		IF SwitchIO.xLiftCylinderExtendInit THEN
		  	IF SwitchIO.xLiftCylinderRetractDetect THEN
		  		iStep:=4;
		  	END_IF;
		  	ELSE
		  	IF SwitchIO.xLiftCylinderExtendDetect THEN
				iStep:=4; 
		  	END_IF;
		END_IF;
		3:(*放行*)	
		ConveyorExitIO.iProductCategory:=ConveyorEntryIO.iProductCategory;
		ConveyorExitIO.iTaskID:=ConveyorEntryIO.iTaskID;
		ConveyorExitIO.diDesConveyor:=ConveyorEntryIO.diDesConveyor;
		SwitchIO.xExitBarCylinderRetract:=1;
		ConveyorExitIO.xPutInto:=0;
		iStep:=4;
		4:(*下料*)
		(*通过出料传输线下料*)
		IF SwitchIO.xExitEnable  AND m_xExitBarDelay AND NOT SwitchIO.xExitBarCylinderRetract  THEN		  
		  	ConveyorExitIO.xUnload:=1;
			ELSE
		  	ConveyorExitIO.xUnload:=0;
		END_IF;	
		(*通过进料传输线下料*)
		IF SwitchIO.xExitEnable  AND m_xExitBarDelay  AND SwitchIO.xExitBarCylinderRetract THEN		  
		  	ConveyorEntryIO.xUnload:=1;
			ELSE
		  	ConveyorEntryIO.xUnload:=0;
		END_IF;			    	
		IF (ConveyorExitIO.xEmpty OR ConveyorEntryIO.xEmpty) AND m_xExitBarDelay  THEN
		  	ConveyorExitIO.xPutInto:=1;
		  	ConveyorEntryIO.xPutInto:=1;
			iStep:=0; 
		END_IF;
	END_CASE;
	m_tonLiftCylinderDelay(IN:=NOT ConveyorEntryIO.xEmpty AND iStep=1 ,PT:= T#1S ,Q:= m_xLiftCylinderDelay ,ET:=m_tLiftCylinderDelay );
	m_tonExitBarDelay(IN:=iStep=4 ,PT:= T#1s ,Q:= m_xExitBarDelay ,ET:= m_tExitBarDelay);
END_IF;
(*复位程序*)
IF (g_xResetSingle AND  (g_diDeviceIDSelect=ConveyorEntryIO.diDeviceID OR g_diDeviceIDSelect=ConveyorExitIO.diDeviceID))
	OR LDP(TRUE,SwitchIO.xLiftCylinderExtendInit) 
	OR LDF(TRUE,SwitchIO.xLiftCylinderExtendInit) 
	OR LDP(TRUE,SwitchIO.xPutInto)  THEN
	ConveyorEntryIO.xPutInto:=1;
	ConveyorExitIO.xPutInto:=1;
	iStep:=0;
END_IF;

IF g_xManual  THEN
	iStep:=0;
	ConveyorEntryIO.xLoad:=0;
    ConveyorEntryIO.xUnload:=0;
	ConveyorEntryIO.xPutInto:=0;
	ConveyorExitIO.xLoad:=0;
	ConveyorExitIo.xUnload:=0;
	ConveyorExitIO.xPutInto:=0;
	SwitchIO.xEntryBarCylinderRetract:=0;
	SwitchIO.xExitBarCylinderRetract:=0;
	IF SwitchIO.xEntryBarCylinderRetractButton THEN
		SwitchIO.xEntryBarCylinderRetract:=1;
		ELSE
		SwitchIO.xEntryBarCylinderRetract:=0;
	END_IF;
	IF SwitchIO.xExitBarCylinderRetractButton THEN
		SwitchIO.xExitBarCylinderRetract:=1;
		ELSE
		SwitchIO.xExitBarCylinderRetract:=0;
	END_IF;
	IF SwitchIO.xLiftCylinderExtendButton AND NOT SwitchIO.xLiftCylinderRetractButton THEN
		SwitchIO.xLiftCylinderExtend:=1;
		SwitchIO.xLiftCylinderRetract:=0;
	END_IF;
	IF NOT SwitchIO.xLiftCylinderExtendButton AND  SwitchIO.xLiftCylinderRetractButton THEN
		SwitchIO.xLiftCylinderExtend:=0;
		SwitchIO.xLiftCylinderRetract:=1;
	END_IF;		 
END_IF;
(*气缸超时报警*)
m_tonCylinderOvertime(IN:= (SwitchIO.xLiftCylinderExtend AND NOT SwitchIO.xLiftCylinderExtendDetect) 
OR  (SwitchIO.xLiftCylinderRetract AND NOT SwitchIO.xLiftCylinderRetractDetect) ,
PT:= SwitchIO.tSetOvertime ,Q:= SwitchIO.xOvertimeAlarm ,ET:= m_tCylinderOvertimeCurrent );
END_FUNCTION_BLOCK

PROGRAM TCP
VAR
  m_ton1ReceiveHeartbeat : TON;
  m_t1RecHeartbeatCurrentTime : TIME;
  m_tonAutoClose : TON;
  m_xAutoClose : BOOL;
  m_tAutoCloseCurrentTime : TIME;
  m_tonReconnect : TON;
  m_ton5ReceiveHeartbeat : TON;
  m_t5RecHeartbeatCurrentTime : TIME;
  m_tonAutoClose1 : TON;
  m_xAutoClose1 : BOOL;
  m_tAutoCloseCurrentTime1 : TIME;
  m_xReconnect : BOOL;
  m_tReconnectCurrentTime : TIME;
  m_tonReconnect1 : TON;
  m_xReconnect1 : BOOL;
  m_tReconnectCurrentTime1 : TIME;
  m_iScanTime : INT;  (* 扫码成功所需时间 *)
  m_iScanTimeMax : INT;  (* 扫码成功所需最长时间 *)
END_VAR
D200:=2;
m_tonReconnect(IN:= NOT SD1282.0 AND NOT SD1284.0 AND NOT m_xReconnect,PT:=T#5s  ,Q:=m_xReconnect ,ET:=m_tReconnectCurrentTime);
SP_SOCOPEN(m_xReconnect  AND SD1288.A , "U0", K1 , D100 , M100);
SP_SOCSND( SM412 AND SD1282.0 , "U0" , K1 , D110, D200, M102 );
SP_SOCRCV( SD1282.0 AND SD1286.0 AND NOT M104 , "U0" , K1, D120 , D400 ,M104 );
m_tonAutoClose(IN:= SD1284.0 AND NOT SD1282.0 ,PT:=T#5s,Q:=m_xAutoClose ,ET:= m_tAutoCloseCurrentTime );
SP_SOCCLOSE( LDF(TRUE,SD1282.0) OR m_xAutoClose  , "U0" , K1, D130, M106 );
D201.F:=SM413;
m_ton1ReceiveHeartbeat(IN:=NOT LDP(TRUE, D401.F) ,PT:= t#5S ,Q:= g_xTcpFailed ,ET:= m_t1RecHeartbeatCurrentTime);
IF g_xTcpFailed THEN
	M104:=SM413;(*通讯失败有可能是接收模块没动作，重启接收模块*)
	D400:=0;
	D401:=0;
END_IF;

(*测试一下通信恢复功能*)
IF  LDP(TRUE,g_xTcpFailed) THEN
	SD1284.0:=SM414;
	SD414:=20;
END_IF;	

D220:=4;
D221:=H54;(*16进制的54转成ASCII码就是T，扫码枪设定的扫码触发条件*)
m_tonReconnect1(IN:= NOT SD1282.4 AND NOT SD1284.4 AND NOT m_xReconnect1 ,PT:=T#5s  ,Q:=m_xReconnect1 ,ET:=m_tReconnectCurrentTime1);
SP_SOCOPEN(m_xReconnect1  AND SD1288.A , "U0", K5 , D140, M108);
SP_SOCSND( LDP(TRUE,g_xScan (*AND NOT g_xScanOvertime*)) AND SD1282.4 , "U0" , K5 , D150, D220, M110);
SP_SOCRCV( SD1282.4 AND SD1286.4 AND NOT M112, "U0" , K5, D160, g_iBatteryInformation[0],M112);
m_tonAutoClose1(IN:= SD1284.4 AND NOT SD1282.4 ,PT:=T#5s,Q:=m_xAutoClose1 ,ET:= m_tAutoCloseCurrentTime1 );
SP_SOCCLOSE( LDF(TRUE,SD1282.4) OR m_xAutoClose1  , "U0" , K5, D170, M114);
(*
IF g_xScan AND g_iBatteryInformation[0]=0 AND ldp(TRUE,SM410) THEN
	MOV( m_iScanTime>m_iScanTimeMax, m_iScanTime , m_iScanTimeMax );
	m_iScanTime:=m_iScanTime+1;
ELSIF NOT g_xScan THEN	*)(*这里统计一下从我发扫码信号，到他扫出结果，所需最长时间*)(*
	g_iBatteryInformation[0]:=0;
	m_iScanTime:=0;
END_IF;	*)
END_PROGRAM

FUNCTION_BLOCK UConveyor
VAR
  iStep : INT;
END_VAR
VAR_IN_OUT
  ConveyorIOLeft : ConveyorIO;  (* U的左半边 *)
  ConveyorIORight : ConveyorIO;  (* U的右半边 *)
  ConveyorIODown : ConveyorIO;  (* U的下边一横 *)
  UConveyorIO : UConveyorIO;  (* 顶升,阻挡 *)
END_VAR
VAR
  m_xInitial : BOOL;
  m_tonCylinderOvertime : TON;  (* 气缸超时报警定时器 *)
  m_tCylinderOvertimeCurrent : TIME;
  m_tonExitBarDelay : TON;  (* 退出阻挡器延时 *)
  m_tExitBarDelay : TIME;
  m_xExitBarDelay : BOOL;
  m_TonStep0 : TON;  (* Step为0延时 *)
  m_xStep0 : BOOL;  (* Step为0延时 *)
  m_tStep0 : TIME;  (* Step为0延时 *)
END_VAR
(*                                                                                                          
初始化中增加气缸复位，气缸位置有BUG
//*)
IF NOT m_xInitial THEN
	UConveyorIO.tSetOvertime:=T#5s;
	UConveyorIO.xExitEnable1:=1;
	UConveyorIO.xExitEnable2:=1;
	UConveyorIO.xExitEnable3:=1;
	m_xInitial:=1;
END_IF;
(*外部不用写ConveyorDown的开关，会自己根据来料的产品信息判断停哪个光电*)
IF UConveyorIO.iTask=1 AND ConveyorIODown.diDesConveyorIn=ConveyorIOLeft.diDeviceID THEN
	ConveyorIODown.xCWPresent:=ConveyorIOLeft.xCCWPresent;
ELSIF UConveyorIO.iTask=1 AND ConveyorIODown.diDesConveyorIn=ConveyorIORight.diDeviceID THEN
	ConveyorIODown.xCWPresent:=ConveyorIORight.xCCWPresent;
ELSE
	ConveyorIODown.xCWPresent:=ConveyorIOLeft.xCCWPresent OR ConveyorIORight.xCCWPresent;
END_IF;
(*这里判断什么时候直接放行，左右都不需要，也不是0，就放走*)
IF  NOT(ConveyorIODown.diDesConveyor=ConveyorIOLeft.diDeviceID 
		OR  ConveyorIODown.diDesConveyor=ConveyorIORight.diDeviceID 
		OR ConveyorIODown.diDesConveyor=0) THEN
	UConveyorIO.xPassEnable:=1;
ELSE
	UConveyorIO.xPassEnable:=0;
END_IF;	
IF g_xAuto THEN	
(*	//加个Step为0的延时，防止扫描周期的影响*)
	m_TonStep0(IN:= iStep=0 ,PT:= t#100ms ,Q:= m_xStep0 ,ET:= m_tStep0 );
	(*//这个是留给阻挡动作的时间*)
	m_tonExitBarDelay(IN:=iStep=4 ,PT:= T#1s ,Q:= m_xExitBarDelay ,ET:= m_tExitBarDelay);
CASE UConveyorIO.iTask OF(*这个Task做抢占，可做LastTask保护*)
0:(*各种初始化，能自动去3*)
	ConveyorIODown.xLoad:=0;
	ConveyorIOleft.xLoad:=0;
	ConveyorIORight.xLoad:=0;
	ConveyorIODown.xUnload:=0;
	ConveyorIOLeft.xUnload:=0;
	ConveyorIORight.xUnload:=0;
	ConveyorIODown.xPutInto:=0;
	ConveyorIOLeft.xPutInto:=0;
	ConveyorIORight.xPutInto:=0;	
	UConveyorIO.xExitBarCylinderRetract1:=0;
	UConveyorIO.xExitBarCylinderRetract2:=0;	
	UConveyorIO.xLiftCylinderRetract1:=1;
	UConveyorIO.xLiftCylinderRetract2:=1;
	UConveyorIO.xLiftCylinderExtend1:=0;
	UConveyorIO.xLiftCylinderExtend2:=0;
1:(*上料*)
	CASE iStep OF
	0:(*各种初始化，能自动去3*)
		ConveyorIODown.xLoad:=0;
		ConveyorIOleft.xLoad:=0;
		ConveyorIORight.xLoad:=0;
		ConveyorIODown.xUnload:=0;
		ConveyorIOLeft.xUnload:=0;
		ConveyorIORight.xUnload:=0;
		UConveyorIO.xExitBarCylinderRetract1:=0;
		UConveyorIO.xExitBarCylinderRetract2:=0;
		UConveyorIO.xBatteryError:=0;
		ConveyorIODown.xPutInto:=0;
		ConveyorIOLeft.xPutInto:=0;
		ConveyorIORight.xPutInto:=0;	
	(*	//根据是否有料判断去1还是3，但会等一个延时*)
		IF m_xStep0 AND  ConveyorIODown.xEmpty THEN
			iStep:=1;
		ELSIF m_xStep0 AND NOT ConveyorIODown.xEmpty THEN
			iStep:=3;
		END_IF;	
	1:(*顶升初始化，等load*)
		(*//左顶升*)
		IF UConveyorIO.xLiftCylinderExtendInit1 THEN
			UConveyorIO.xLiftCylinderExtend1:=1;
			UConveyorIO.xLiftCylinderRetract1:=0;
		ELSE
			UConveyorIO.xLiftCylinderExtend1:=0;
			UConveyorIO.xLiftCylinderRetract1:=1;
		END_IF;
	(*	//右顶升*)
		IF UConveyorIO.xLiftCylinderExtendInit2 THEN
			UConveyorIO.xLiftCylinderExtend2:=1;
			UConveyorIO.xLiftCylinderRetract2:=0;
			ELSE
			UConveyorIO.xLiftCylinderExtend2:=0;
			UConveyorIO.xLiftCylinderRetract2:=1;
		END_IF;
		(*//顶升到位，等上料信号*)
		IF 	((UConveyorIO.xLiftCylinderExtendInit1 AND UConveyorIO.xLiftCylinderExtendDetect1)
				OR (NOT UConveyorIO.xLiftCylinderExtendInit1 AND UConveyorIO.xLiftCylinderRetractDetect1))
			AND	((UConveyorIO.xLiftCylinderExtendInit2 AND UConveyorIO.xLiftCylinderExtendDetect2)
		   		OR (NOT UConveyorIO.xLiftCylinderExtendInit2 AND UConveyorIO.xLiftCylinderRetractDetect2))		
			AND	UConveyorIO.xEntryEnable1 THEN(*有上料请求1*)
		   	ConveyorIODown.xLoad:=1;
			iStep:=2;
		END_IF;
	2:(*Load完成*)
		(*去右臂时才需要阻挡1放行,其他情况阻挡1挡住*)
		UConveyorIO.xExitBarCylinderRetract1:=ConveyorIODown.diDesConveyorIn=ConveyorIORight.diDeviceID;
		IF NOT ConveyorIODown.xEmpty THEN
			ConveyorIODown.xLoad:=0;
			ConveyorIOLeft.xPutInto:=1;
			ConveyorIOright.xPutInto:=1;
			istep:=3;
		END_IF;
	3:(*顶升等Unload，这里等有了ExitEnable再顶升，因为可能有地方需要允许了再升降，比如倍速链*)
		(*//电池检测保护，防止把带电池的料框送进去了*)
		IF (ConveyorIODown.diDesConveyor=ConveyorIOLeft.diDeviceID OR ConveyorIODown.diDesConveyor=ConveyorIORight.diDeviceID)
			AND	(UConveyorIO.xBatteryDetect1 OR UConveyorIO.xBatteryDetect2)(*在下面时检测*)
			AND UConveyorIO.xLiftCylinderRetractDetect1 AND UConveyorIO.xLiftCylinderRetractDetect2 THEN
			UConveyorIO.xBatteryError:=1;
		END_IF;	
		(*//左侧顶升控制*)
		IF (ConveyorIODown.diDesConveyor=ConveyorIOLeft.diDeviceID AND UConveyorIO.xExitEnable2 AND NOT UConveyorIO.xBatteryError)THEN
			IF UConveyorIO.xLiftCylinderExtendInit1 THEN
				UConveyorIO.xLiftCylinderExtend1:=0;
				UConveyorIO.xLiftCylinderRetract1:=1;
			ELSE
				UConveyorIO.xLiftCylinderExtend1:=1;
				UConveyorIO.xLiftCylinderRetract1:=0;
			END_IF;
			IF(NOT UConveyorIO.xLiftCylinderExtendInit1 AND UConveyorIO.xLiftCylinderExtendDetect1)
				OR (UConveyorIO.xLiftCylinderExtendInit1 AND UConveyorIO.xLiftCylinderRetractDetect1)THEN
				ConveyorIOLeft.xPutInto:=0;
				ConveyorIOright.xPutInto:=0;
				iStep:=4;
			END_IF;
		END_IF;	
		(*//右侧顶升控制*)
		IF (ConveyorIODown.diDesConveyor=ConveyorIORight.diDeviceID AND UConveyorIO.xExitEnable3 AND NOT UConveyorIO.xBatteryError)THEN
			IF UConveyorIO.xLiftCylinderExtendInit2 THEN
				UConveyorIO.xLiftCylinderExtend2:=0;
				UConveyorIO.xLiftCylinderRetract2:=1;
			ELSE
				UConveyorIO.xLiftCylinderExtend2:=1;
				UConveyorIO.xLiftCylinderRetract2:=0;
			END_IF;
			IF(NOT UConveyorIO.xLiftCylinderExtendInit2 AND UConveyorIO.xLiftCylinderExtendDetect2)
				OR (UConveyorIO.xLiftCylinderExtendInit2 AND UConveyorIO.xLiftCylinderRetractDetect2) THEN
				ConveyorIOLeft.xPutInto:=0;
				ConveyorIOright.xPutInto:=0;
				iStep:=4;
			END_IF;
		END_IF;	
	(*	//直接放行控制*)
		IF UConveyorIO.xPassEnable AND UConveyorIO.xExitEnable1 AND NOT UConveyorIO.xBatteryError THEN
			IF UConveyorIO.xLiftCylinderExtendInit1 THEN
				UConveyorIO.xLiftCylinderExtend1:=1;
				UConveyorIO.xLiftCylinderRetract1:=0;
			ELSE
				UConveyorIO.xLiftCylinderExtend1:=0;
				UConveyorIO.xLiftCylinderRetract1:=1;
			END_IF;
			IF UConveyorIO.xLiftCylinderExtendInit2 THEN
				UConveyorIO.xLiftCylinderExtend2:=1;
				UConveyorIO.xLiftCylinderRetract2:=0;
			ELSE
				UConveyorIO.xLiftCylinderExtend2:=0;
				UConveyorIO.xLiftCylinderRetract2:=1;
			END_IF;
			IF((UConveyorIO.xLiftCylinderExtendInit1 AND UConveyorIO.xLiftCylinderExtendDetect1)
 OR (NOT UConveyorIO.xLiftCylinderExtendInit1 AND UConveyorIO.xLiftCylinderRetractDetect1))
				AND((UConveyorIO.xLiftCylinderExtendInit2 AND UConveyorIO.xLiftCylinderExtendDetect2)
 OR (NOT UConveyorIO.xLiftCylinderExtendInit2 AND UConveyorIO.xLiftCylinderRetractDetect2))THEN
				UConveyorIO.xExitBarCylinderRetract1:=1;
				UConveyorIO.xExitBarCylinderRetract2:=1;
				ConveyorIOLeft.xPutInto:=0;
				ConveyorIOright.xPutInto:=0;
				iStep:=4;
			END_IF;	
		END_IF;
	4:(*Unload完成，回0*)
			IF ConveyorIODown.diDesConveyor=ConveyorIOLeft.diDeviceID AND UConveyorIO.xExitEnable2 AND m_xExitBarDelay THEN
				ConveyorIOLeft.xUnload:=1;
			ELSIF ConveyorIODown.diDesConveyor=ConveyorIORight.diDeviceID AND UConveyorIO.xExitEnable3 AND m_xExitBarDelay THEN
				ConveyorIORight.xUnload:=1;
			ELSIF UConveyorIO.xPassEnable AND UConveyorIO.xExitEnable1 AND m_xExitBarDelay THEN
				ConveyorIODown.xUnload:=1;
			ELSE
				ConveyorIODown.xUnload:=0;
				ConveyorIOLeft.xUnload:=0;
				ConveyorIORight.xUnload:=0;
			END_IF;	
		IF ( (ConveyorIODown.diDesConveyor=ConveyorIOLeft.diDeviceID  AND LDF(TRUE,UConveyorIO.xExitEnable2))
		  OR(ConveyorIODown.diDesConveyor=ConveyorIORight.diDeviceID AND LDF(TRUE,UConveyorIO.xExitEnable3))
		  OR(UConveyorIO.xPassEnable AND LDF(TRUE,UConveyorIO.xExitEnable1)) )AND m_xExitBarDelay  THEN
			ConveyorIODown.xUnload:=0;
			ConveyorIOLeft.xUnload:=0;
			ConveyorIORight.xUnload:=0;
			ConveyorIODown.xPutInto:=1;
			ConveyorIOLeft.xPutInto:=1;
			ConveyorIORight.xPutInto:=1;
			UConveyorIO.xExitBarCylinderRetract1:=0;
			UConveyorIO.xExitBarCylinderRetract2:=0;
			iStep:=0;
		END_IF;
	END_CASE;
2:(*左下料*)
	CASE iStep OF
	0:(*各种初始化，能自动去3*)
		ConveyorIODown.xLoad:=0;
		ConveyorIOleft.xLoad:=0;
		ConveyorIORight.xLoad:=0;
		ConveyorIODown.xUnload:=0;
		ConveyorIOLeft.xUnload:=0;
		ConveyorIORight.xUnload:=0;
		UConveyorIO.xBatteryError:=0;
		UConveyorIO.xExitBarCylinderRetract1:=0;
		UConveyorIO.xExitBarCylinderRetract2:=0;
		ConveyorIODown.xPutInto:=0;
		ConveyorIOLeft.xPutInto:=0;
		ConveyorIORight.xPutInto:=0;
		IF m_xStep0 AND  ConveyorIODown.xEmpty THEN
			iStep:=1;
		ELSIF m_xStep0 AND NOT ConveyorIODown.xEmpty THEN
			iStep:=3;
		END_IF;	
	1:(*左顶升动作，等load*)
		IF UConveyorIO.xLiftCylinderExtendInit1 THEN
			UConveyorIO.xLiftCylinderExtend1:=0;
			UConveyorIO.xLiftCylinderRetract1:=1;
			ELSE
			UConveyorIO.xLiftCylinderExtend1:=1;
			UConveyorIO.xLiftCylinderRetract1:=0;
		END_IF;
		IF ((NOT UConveyorIO.xLiftCylinderExtendInit1 AND UConveyorIO.xLiftCylinderExtendDetect1)
			OR ( UConveyorIO.xLiftCylinderExtendInit1 AND UConveyorIO.xLiftCylinderRetractDetect1))
			AND UConveyorIO.xEntryEnable2 THEN(*有上料请求1*)
		   	ConveyorIOLeft.xLoad:=1;
			iStep:=2;
		END_IF;
	2:(*Load完成*)
		IF NOT ConveyorIOLeft.xEmpty THEN
			ConveyorIOLeft.xLoad:=0;
			ConveyorIODown.xPutInto:=1;
			ConveyorIODown.diDesConveyor:=ConveyorIOLeft.diDesConveyor;
			istep:=3;
		END_IF;
	3:(*顶升等Unload，这里等有了ExitEnable再顶升，因为可能有地方需要允许了再升降，比如倍速链*)
		UConveyorIO.xExitBarCylinderRetract1:=1;
		UConveyorIO.xExitBarCylinderRetract2:=1;
		IF  UConveyorIO.xExitEnable1 THEN
			IF UConveyorIO.xLiftCylinderExtendInit1 THEN
				UConveyorIO.xLiftCylinderExtend1:=1;
				UConveyorIO.xLiftCylinderRetract1:=0;
			ELSE
				UConveyorIO.xLiftCylinderExtend1:=0;
				UConveyorIO.xLiftCylinderRetract1:=1;
			END_IF;
			IF(( UConveyorIO.xLiftCylinderExtendInit1 AND UConveyorIO.xLiftCylinderExtendDetect1)
				OR (NOT UConveyorIO.xLiftCylinderExtendInit1 AND UConveyorIO.xLiftCylinderRetractDetect1))THEN
				ConveyorIODown.xPutInto:=0;
				iStep:=4;
			END_IF;	
		END_IF;
	4:(*Unload完成，回0*)
		IF  UConveyorIO.xExitEnable1 AND m_xExitBarDelay THEN
			ConveyorIODown.xUnload:=1;
		ELSE
			ConveyorIODown.xUnload:=0;
		END_IF;	
		IF NOT UConveyorIO.xExitEnable1 AND m_xExitBarDelay   THEN
			ConveyorIODown.xUnload:=0;
			ConveyorIOLeft.xUnload:=0;
			ConveyorIORight.xUnload:=0;
			ConveyorIODown.xPutInto:=1;
			ConveyorIOLeft.xPutInto:=1;
			ConveyorIORight.xPutInto:=1;
			UConveyorIO.xExitBarCylinderRetract1:=0;
			UConveyorIO.xExitBarCylinderRetract2:=0;
			iStep:=0;
		END_IF;
	END_CASE;
3:(*上料到出口*)
	CASE iStep OF
	0:(*各种初始化，能自动去3*)
		ConveyorIODown.xLoad:=0;
		ConveyorIOleft.xLoad:=0;
		ConveyorIORight.xLoad:=0;
		ConveyorIODown.xUnload:=0;
		ConveyorIOLeft.xUnload:=0;
		ConveyorIORight.xUnload:=0;
		UConveyorIO.xBatteryError:=0;
		UConveyorIO.xExitBarCylinderRetract1:=0;
		UConveyorIO.xExitBarCylinderRetract2:=0;
		ConveyorIODown.xPutInto:=0;
		ConveyorIOLeft.xPutInto:=0;
		ConveyorIORight.xPutInto:=0;
		IF m_xStep0 AND  ConveyorIODown.xEmpty THEN
			iStep:=1;
		ELSIF m_xStep0 AND NOT ConveyorIODown.xEmpty THEN
			iStep:=3;
		END_IF;	
	1:(*右顶升动作，等load*)
		IF UConveyorIO.xLiftCylinderExtendInit2 THEN
			UConveyorIO.xLiftCylinderExtend2:=0;
			UConveyorIO.xLiftCylinderRetract2:=1;
		ELSE
			UConveyorIO.xLiftCylinderExtend2:=1;
			UConveyorIO.xLiftCylinderRetract2:=0;
		END_IF;
		IF ((NOT UConveyorIO.xLiftCylinderExtendInit2 AND UConveyorIO.xLiftCylinderExtendDetect2)
			OR ( UConveyorIO.xLiftCylinderExtendInit2 AND UConveyorIO.xLiftCylinderRetractDetect2))
			AND UConveyorIO.xEntryEnable3 THEN(*有上料请求1*)
		   	ConveyorIORight.xLoad:=1;
			iStep:=2;
		END_IF;
	2:(*Load完成*)
		IF NOT ConveyorIORight.xEmpty THEN
			ConveyorIORight.xLoad:=0;
			ConveyorIODown.diDesConveyor:=ConveyorIORight.diDesConveyor;
			ConveyorIODown.xPutInto:=1;
			istep:=3;
		END_IF;
	3:(*顶升恢复等Unload，这里等有了ExitEnable再顶升，因为可能有地方需要允许了再升降，比如倍速链*)
		UConveyorIO.xExitBarCylinderRetract2:=1;
		IF  UConveyorIO.xExitEnable1 THEN(**)
			IF UConveyorIO.xLiftCylinderExtendInit2 THEN
				UConveyorIO.xLiftCylinderExtend2:=1;
				UConveyorIO.xLiftCylinderRetract2:=0;
			ELSE
				UConveyorIO.xLiftCylinderExtend2:=0;
				UConveyorIO.xLiftCylinderRetract2:=1;
			END_IF;
		END_IF;
		IF UConveyorIO.xExitEnable1 THEN(**)
			IF(( UConveyorIO.xLiftCylinderExtendInit2 AND UConveyorIO.xLiftCylinderExtendDetect2)
				OR (NOT UConveyorIO.xLiftCylinderExtendInit2 AND UConveyorIO.xLiftCylinderRetractDetect2))THEN
				ConveyorIODown.xPutInto:=0;
				iStep:=4;
			END_IF;	
		END_IF;
	4:(*Unload完成，回0*)
		IF  UConveyorIO.xExitEnable1 AND m_xExitBarDelay THEN
			ConveyorIODown.xUnload:=1;
		ELSE
			ConveyorIODown.xUnload:=0;
		END_IF;	
		IF NOT UConveyorIO.xExitEnable1 AND m_xExitBarDelay  THEN
			ConveyorIODown.xUnload:=0;
			ConveyorIOLeft.xUnload:=0;
			ConveyorIORight.xUnload:=0;
			ConveyorIODown.xPutInto:=1;
			ConveyorIOLeft.xPutInto:=1;
			ConveyorIORight.xPutInto:=1;
			UConveyorIO.xExitBarCylinderRetract1:=0;
			UConveyorIO.xExitBarCylinderRetract2:=0;
			iStep:=0;
		END_IF;
	END_CASE;
END_CASE;(*iTask*)
END_IF;(*g_xAuto那个IF*)
(*复位程序*)
IF (g_xResetSingle AND  (g_diDeviceIDSelect=ConveyorIOLeft.diDeviceID 
 	 OR g_diDeviceIDSelect=ConveyorIORight.diDeviceID
 	 OR g_diDeviceIDSelect=ConveyorIODown.diDeviceID))
	OR LDP(TRUE,UConveyorIO.xLiftCylinderExtendInit1) 
	OR LDF(TRUE,UConveyorIO.xLiftCylinderExtendInit1) 
	OR LDP(TRUE,UConveyorIO.xPutInto)  THEN
	ConveyorIODown.xPutInto:=1;
	ConveyorIOLeft.xPutInto:=1;
	ConveyorIORight.xPutInto:=1;
	iStep:=0;
END_IF;
(*手动*)
IF g_xManual  THEN
	iStep:=0;
	ConveyorIODown.xLoad:=0;
	ConveyorIOleft.xLoad:=0;
	ConveyorIORight.xLoad:=0;
	ConveyorIODown.xUnload:=0;
	ConveyorIOLeft.xUnload:=0;
	ConveyorIORight.xUnload:=0;
	ConveyorIODown.xPutInto:=0;
	ConveyorIOLeft.xPutInto:=0;
	ConveyorIORight.xPutInto:=0;
	UConveyorIO.xBatteryError:=0;
	UConveyorIO.xLiftCylinderExtend1:=UConveyorIO.xLiftCylinderExtendButton1 AND NOT UConveyorIO.xLiftCylinderRetractButton1;
	UConveyorIO.xLiftCylinderRetract1:=UConveyorIO.xLiftCylinderRetractButton1 AND NOT UConveyorIO.xLiftCylinderExtendButton1;
	UConveyorIO.xLiftCylinderExtend2:=UConveyorIO.xLiftCylinderExtendButton2 AND NOT UConveyorIO.xLiftCylinderRetractButton2;
	UConveyorIO.xLiftCylinderRetract2:=UConveyorIO.xLiftCylinderRetractButton2 AND NOT UConveyorIO.xLiftCylinderExtendButton2;
	UConveyorIO.xExitBarCylinderRetract1:=UConveyorIO.xExitBarCylinderRetractButton1;
	UConveyorIO.xExitBarCylinderRetract2:=UConveyorIO.xExitBarCylinderRetractButton2;
END_IF;	
(*气缸超时报警*)
m_tonCylinderOvertime(IN:= (UConveyorIO.xLiftCylinderExtend1 AND NOT UConveyorIO.xLiftCylinderExtendDetect1) 
 		OR  (UConveyorIO.xLiftCylinderRetract1 AND NOT UConveyorIO.xLiftCylinderRetractDetect1)
 		OR	(UConveyorIO.xLiftCylinderExtend2 AND NOT UConveyorIO.xLiftCylinderExtendDetect2) 
 		OR  (UConveyorIO.xLiftCylinderRetract2 AND NOT UConveyorIO.xLiftCylinderRetractDetect2),
 PT:= UConveyorIO.tSetOvertime ,Q:=UConveyorIO.xOvertimeAlarm ,ET:=m_tCylinderOvertimeCurrent );
END_FUNCTION_BLOCK

PROGRAM 批量复制专用

END_PROGRAM

FUNCTION_BLOCK FanucRobot
VAR_IN_OUT
  FanucRobotIO : FanucRobotIO;
END_VAR
VAR
  m_iSNO : INT;
  m_xPNSPass : BOOL;  (* 收到程序号 *)
  m_tonStartDelay : TON;  (* 启动延时 *)
  m_xStartDelay : BOOL;
  m_tStartDelayCurrentTime : TIME;
END_VAR
(***********************************************************
发那科机器人自动启动程序


***********************************************************)

(*无自动状态，示教盒处于本地状态，把各标志位复位*)
IF FanucRobotIO.i_xTPENBL AND NOT g_xAuto THEN
	FanucRobotIO.o_xPNSTROBE:=0;
	FanucRobotIO.o_xCSTOPI:=0;
	FanucRobotIO.o_xPROD_START:=0;
	FanucRobotIO.o_xRESET:=0;
END_IF;
(*远程模式*)
IF g_xAuto THEN
	FanucRobotIO.o_xREMOTE:=1;
	ELSE
	FanucRobotIO.o_xREMOTE:=0;
END_IF;
(*程序启动后复位启动标志位*)
IF FanucRobotIO.i_xPROG_RUN AND FanucRobotIO.i_xBUSY THEN
	FanucRobotIO.i_xCommandStart:=0;
END_IF;
(*示教盒旋清除报警*)
IF ldf(TRUE,FanucRobotIO.i_xTPENBL)THEN
	FanucRobotIO.o_xRESET:=1;
	FanucRobotIO.o_xCSTOPI:=1;
END_IF;
(*启动程序号条件*)
IF FanucRobotIO.i_xSYSRDY 
	AND FanucRobotIO.i_xCMDENBL
	AND FanucRobotIO.i_xCommandStart
	AND NOT FanucRobotIO.i_xPROG_RUN 
	AND NOT FanucRobotIO.i_xBUSY THEN
	FanucRobotIO.o_xRESET:=0;
	FanucRobotIO.o_xCSTOPI:=0;
	IF FanucRobotIO.i_iMotionNumber <> 0 (*只要动作编号不为0，就给他信号*)
		AND NOT FanucRobotIO.o_xPNSTROBE THEN
		FanucRobotIO.o_xPNSTROBE:=1;
		FanucRobotIO.o_xPROD_START:=1;
		FanucRobotIO.o_iPNS:=FanucRobotIO.i_iMotionNumber;(*并把任务号传给他*)
	END_IF;
	(*程序号校验*)
	IF FanucRobotIO.i_xSNACK THEN(*数据传回之后再校验*)
		m_iSNO:=BITARR_TO_INT(FanucRobotIO.i_arrxSNO[0] , 8 );
		IF m_iSNO=FanucRobotIO.o_iPNS THEN
			m_xPNSPass:=1;(*校验成功,等100MS复位Start信号*)
			FanucRobotIO.o_xPNSTROBE:=0;
		ELSE
			FanucRobotIO.o_xPNSFailed:=1;(*校验失败*)
			FanucRobotIO.o_xPROD_START:=0;(*立刻复位，不生成任务*)
		END_IF;
	END_IF;
END_IF;
m_tonStartDelay(IN:= m_xPNSPass ,PT:= T#100ms ,Q:= m_xStartDelay ,ET:=m_tStartDelayCurrentTime );
IF m_xStartDelay THEN
	FanucRobotIO.o_xPROD_START:=0;
	FanucRobotIO.i_xCommandStart:=0;
	m_xPNSPass:=0;
END_IF;
END_FUNCTION_BLOCK

FUNCTION_BLOCK ConveyorCommunication
VAR_IN_OUT
  ConveyorIO : ConveyorIO;
  CommunicationIO : CommunicationIO;
END_VAR
VAR_OUTPUT
  o_iErrorNub : INT;  (* 错误代码 *)
END_VAR
VAR
  o_xReqSuccess : BOOL;  (* 请求成功 *)
END_VAR
(********************************************************************************)
(*
DB1区(PC->PLC)15个字		
"字(16位）序号
(从1开始)"			功能描述  	具体参数解释
1 请求确认	"  1：复位
				   				2：读码(入库申请）成功
				   				3：取放货完成 
   			4：旋转
   			5：不旋转
   			101：条码空
   			102：条码规则校验失败
   			103：步号校验失败
   			104：无库位可用 
"
2	预留	
3	预留	
4	预留	
5	预留	
6	读写标志位	"  				1：写入数据
   			2：读数据完成"
7	任务处理标志	"  				１：复位
   			２：完成"
8	命令字	"
   			21-送出（任务起点与终点不同，即向下一台输送机移载）
   			22：叠盘
"
9	任务号	"   1~65535唯一任务标识"
10	目标设备号   只有送出任务才有效
11		
12	筐码后4位	
				

DB2区(PLC->PC)15个字			
"字(16位）序号
(从1开始)"	功能描述	具体参数解释	
1	请求状态	"１：复位
２：请求"	实时状态，没有时序交互
2	强制入库(预留）	"１：复位
２：强制入库"	
3	预留(叠盘数量）	只对叠盘工位有效	
4	预留		
5			
6	读写标志位	"1：写入数据
2：读数据完成"	"有交互
时序"
7	设备状态	"1:空闲
2：工作中
3:任务完成（只有目标设备才会报任务完成）
４：故障"	
8	任务号	1~65535唯一任务标识，当输送任务执行完成后，将PC下发的任务号上报	
9	筐码后4位		
10	预留		
11			
			





2018.8.3 YAO 1.0
*)
(********************************************************************************)
(*//请求状态*)
IF ConveyorIO.xEmpty THEN
	CommunicationIO.o_iRequestPLCPC:=1;
	ELSE
	CommunicationIO.o_iRequestPLCPC:=2;
END_IF;
(*//请求确认*)
CASE CommunicationIO.i_iResponsPCPLC OF 
	0:;
	1:;(*//复位*)
	2:(*//读码（入库申请）成功*)
	o_xReqSuccess:=1;
	3:(*//取放货完成*)
	ConveyorIO.xPutInto:=1; 
	4:(*//旋转*)
	;
	5:(*//不旋转*)
	;
	101:(*//条码空*)
	o_iErrorNub:=101;
	102:(*//条码规则检验失败*)
	o_iErrorNub:=102;
	103:(*//步号校验失败*)
	o_iErrorNub:=103;
	104:(*//无库位可用*)
	o_iErrorNub:=104;
END_CASE;
IF CommunicationIO.i_iResponsPCPLC <> 3 THEN
	ConveyorIO.xPutInto:=0;
END_IF;
IF CommunicationIO.i_iResponsPCPLC <> 2 THEN
	o_xReqSuccess:=0;
END_IF;
IF CommunicationIO.i_iResponsPCPLC < 100 THEN
	o_iErrorNub:=0;
END_IF;

(*//读写标志位写入数据*)
IF LDP(TRUE,CommunicationIO.i_iReadWriteFlagPCPLC = 1) THEN
	ConveyorIO.iTaskID := CommunicationIO.i_iTaskIDPCPLC;
	ConveyorIO.diDesConveyor := CommunicationIO.i_diDestinationDevicePCPLC;
	ConveyorIO.iProductCategory := CommunicationIO.i_iProductIDPCPLC;
END_IF;
(*//数据校验，并返回握手信号*)
IF CommunicationIO.i_iReadWriteFlagPCPLC = 1 
	AND ConveyorIO.iTaskID<>0
	AND ConveyorIO.diDesConveyor<>0 
	AND ConveyorIO.iProductCategory<>0 
	THEN
	CommunicationIO.o_iReadWriteFlagPLCPC:=2;
	ELSE
	CommunicationIO.o_iReadWriteFlagPLCPC:=1;
END_IF;
(*//数据校验*)
IF CommunicationIO.i_iReadWriteFlagPCPLC = 1 
	AND (ConveyorIO.iTaskID<>0
	OR ConveyorIO.diDesConveyor<>0 
	OR ConveyorIO.iProductCategory<>0) 
	THEN
	o_iErrorNub:=50;(*//任务数据不完整*)
END_IF;
(*//设备状态*)
IF ConveyorIO.diDesConveyor = ConveyorIO.diDeviceID AND NOT ConveyorIO.xEmpty THEN(*//目标地址=当前地址*)
	CommunicationIO.o_iDeviceStatusPLCPC:=3;(*//任务完成*)
	CommunicationIO.o_iProductIDPLCPC:=ConveyorIO.iProductCategory;(*//条码号上传*)
	CommunicationIO.o_iTaskIDPLCPC:=ConveyorIO.iTaskID;(*//任务号上传*)
	ELSIF ConveyorIO.xBusy THEN
	CommunicationIO.o_iDeviceStatusPLCPC:=2;(*//工作中*)
	ELSIF ConveyorIO.xError THEN
	CommunicationIO.o_iDeviceStatusPLCPC:=4;(*//故障*)
	ELSE
	CommunicationIO.o_iDeviceStatusPLCPC:=1;(*//空闲*)
	CommunicationIO.o_iProductIDPLCPC:=0;(*//条码号复位*)
	CommunicationIO.o_iTaskIDPLCPC:=0;(*//任务号复位*)
END_IF;
END_FUNCTION_BLOCK

FUNCTION_BLOCK PackCommunication
VAR_IN_OUT
  ConveyorIO : ConveyorIO;
  PackCommunicationIO : PackCommunicationIO;
  FanucRobotIO : FanucRobotIO;
END_VAR
VAR_OUTPUT
  o_iErrorNub : INT;
  o_xReqSuccess : BOOL;
END_VAR
VAR
  m_xReqSuccess : BOOL;
  m_iStep : INT;
  m_arrwCode : ARRAY [1..8] OF BatteryCode;
END_VAR
VAR_INPUT
  i_arrxPresentDetect : ARRAY [1..8] OF BOOL;
END_VAR
VAR
  m_iCoordinateX : INT;
  m_iCoordinateY : INT;
  m_arriPresentDetect : ARRAY [1..8] OF INT;
  ii : INT;
END_VAR
VAR CONSTANT
  MAX_ROW : INT := 8;
  MAX_COLUMN : INT := 8;
END_VAR
VAR
  m_xSupplement : BOOL;
END_VAR
VAR CONSTANT
  ROW_TIMES : INT := 1;
  GET_QUANTITY : INT := 8;
END_VAR
VAR
  m_iRowReminder : INT;
  m_xEno : BOOL;
  m_iRowReminderTemp : INT;
END_VAR
(***************************************************************************)
(*
DB1区(PC->PLC)10个字		
"字(16位）序号
(从1开始)"	功能描述	具体参数解释
1	请求确认	"1：复位
2：读码(入库申请）成功
101：条码空
102：条码规则校验失败
103：步号校验失败
"
2	放行	"1：复位
2：完成,放行
3：撤销完成 "
3	单次装载应答	"1：复位
2：允许开始"
4	单次装载处理完成	"1：复位
2：完成
3：电芯为空"
)*
DB2区(PLC->PC)200个字		
"字(16位）序号
(从1开始)"	功能描述	具体参数解释
1	装载请求	"１：复位
２：请求"
2	装载全部完成	"1：复位
2：请求 "
3	单次装载请求	"1：复位
2：请求 "
4	单次装载完成	"1：复位
2：完成"
5	行坐标	从1开始
6	列坐标	从1开始
7	电芯码(15*11=165)	"电芯码24字符，
占12个字，加上预留的每个分配15个字"

顺序执行步骤
0  初始化
1  框码扫码请求
2  单次抓取请求
3  整排抓取
4  补料
5  完成


(***************************************************************************)
m_iRowReminder:= ( m_iCoordinateX-1 MOD GET_QUANTITY )+1;(*//通过位置与抓取数量取余数，判断是否的抓取位置为一排的最后一个*)
CASE m_iStep OF
	0:;(*//初始化*)
	m_iStep:=1;
	1:(*发送框码的扫码请求*)
	IF NOT ConveyorIO.xEmpty AND NOT FanucRobotIO.io_xMutexLock THEN
		PackCommunicationIO.o_iRequestPLCPC:=2;
		ELSE
		PackCommunicationIO.o_iRequestPLCPC:=1;
	END_IF;
	(*//请求确认*)
	CASE PackCommunicationIO.i_iResponsPCPLC OF 
		0:;
		1:;(*//复位*)
		2:(*//读码（入库申请）成功*)
		m_iStep:=2;
		m_xSupplement:=0;
		m_iCoordinateX:=1;(*//框码扫码成功后把坐标改为1,1*)
		m_iCoordinateY:=1;
		FanucRobotIO.io_xMutexLock:=1;
		3:(*//取放货完成*)
		ConveyorIO.xPutInto:=1; 
		4:(*//旋转*)
		;
		5:(*//不旋转*)
		;
		101:(*//条码空*)
		o_iErrorNub:=101;
		m_iStep:=0;
		102:(*//条码规则检验失败*)
		o_iErrorNub:=102;
		m_iStep:=0;
		103:(*//步号校验失败*)
		o_iErrorNub:=103;
		m_iStep:=0;
		104:(*//无库位可用*)
		o_iErrorNub:=104;
		m_iStep:=0;
	END_CASE;
	2:(*//单次抓取请求，分为单次多个产品抓取与补料程序*)
	IF FanucRobotIO.i_xSYSRDY 
		AND NOT FanucRobotIO.i_xBUSY
		AND NOT FanucRobotIO.i_xPROG_RUN
		AND i_arrxPresentDetect[1] 
		AND PackCommunicationIO.i_iSinglePackResponsePCPLC=1 THEN(*//机器人准备就绪、组装下线有料*)
		PackCommunicationIO.o_iSinglePackRequestPLCPC:=2;
	END_IF;
	IF (*LDP(TRUE,PackCommunicationIO.i_iSinglePackResponsePCPLC=2)*) PackCommunicationIO.i_iSinglePackResponsePCPLC=2 THEN(*//请求成功*)
		PackCommunicationIO.o_iSinglePackRequestPLCPC:=1;(*//复位请求*)
		IF m_xSupplement THEN(*//补料标志位，为1进行补料操作，为0进行整排抓取*)
			m_iStep:=4;(*//补料*)
			ELSE
		 	m_iStep:=3;(*//整排抓取*)
			FOR ii:=1 TO GET_QUANTITY BY 1 DO(*//记录哪个位置缺料*)
				IF i_arrxPresentDetect[ii] THEN(*//传感器检测*)
 m_arriPresentDetect[ii]:=0;
 ELSE
 m_arriPresentDetect[ii]:=ii;(*//记录缺料的位置*)
				END_IF;
			END_FOR;
		END_IF;
	END_IF;
	3:  (*//整排抓取*)
	FanucRobotIO.o_iPNS:=10101;(*//步骤号*)
	FanucRobotIO.o_uiOffset_X:=m_iCoordinateX;
	FanucRobotIO.o_uiOffset_Y:=m_iCoordinateY;
	PackCommunicationIO.o_iXCoordinatePLCPC:=m_iCoordinateX;(*//放置位置发送给上位机*)
	PackCommunicationIO.o_iYCoordinatePLCPC:=m_iCoordinateY;	
	IF LDF(TRUE,FanucRobotIO.i_xBUSY OR FanucRobotIO.i_xPROG_RUN) THEN(*//抓取动作完成*)
		FOR ii:=1 TO GET_QUANTITY BY 1 DO (*//判断有无补料信息*)
			IF m_arriPresentDetect[ii]<>0  THEN(*//有补料*)(*//补料不是最后一个的算法*)
				m_iCoordinateX:=m_arriPresentDetect[ii]+((m_iCoordinateX-1)/GET_QUANTITY)*GET_QUANTITY;
				m_xSupplement:=1;
				m_iStep:=2;(*//有补料*)
				EXIT;
			END_IF;			
		END_FOR;
		IF ii=GET_QUANTITY+1  THEN  (*//无补料*)
			m_xSupplement:=0;
			IF m_iCoordinateY = MAX_ROW (*//达到最大列*)
				AND ((m_iCoordinateX-1)/GET_QUANTITY+1=ROW_TIMES) 
				THEN(*//偏移量为最大的值时,排抓取为最后一排*)
				m_iStep:=5;(*//装盘完成*)
				ELSE
				m_iStep:=2;(*//请求下一次装盘*)			
				IF (m_iCoordinateX-1)/GET_QUANTITY+1=ROW_TIMES THEN
 m_iCoordinateX:=1;                                              (*//开始执行下一列*)
 m_iCoordinateY:=m_iCoordinateY+1;
 ELSE
 m_iCoordinateX:=((m_iCoordinateX-1)/GET_QUANTITY+1)*GET_QUANTITY+1;
				END_IF;
			END_IF;
		END_IF;
	END_IF;
	4: (*//补料*)
	FanucRobotIO.o_iPNS:=10102;(*//步骤号*)
	FanucRobotIO.o_uiOffset_X:=m_iCoordinateX;
	FanucRobotIO.o_uiOffset_Y:=m_iCoordinateY;
	PackCommunicationIO.o_iXCoordinatePLCPC:=m_iCoordinateX;(*//放置位置发送给上位机*)
	PackCommunicationIO.o_iYCoordinatePLCPC:=m_iCoordinateY;
	IF LDF(TRUE,FanucRobotIO.i_xBUSY OR FanucRobotIO.i_xPROG_RUN) THEN(*//抓取动作完成*)
		FOR ii:=m_iRowReminder+1 TO GET_QUANTITY BY 1 DO (*//判断有无补料信息*)
			IF m_arriPresentDetect[ii]<>0  THEN(*//有补料*)(*//补料不是最后一个的算法*)
				m_iCoordinateX:=m_arriPresentDetect[ii]+((m_iCoordinateX-1)/GET_QUANTITY)*GET_QUANTITY;
				m_xSupplement:=1;
				m_iStep:=2;(*//有补料*)
				EXIT;
			END_IF;	
		END_FOR;
		IF ii=GET_QUANTITY+1  THEN  (*//无补料*)
			m_xSupplement:=0;
			IF m_iCoordinateY = MAX_ROW (*//达到最大列*)
				AND ((m_iCoordinateX-1)/GET_QUANTITY+1=ROW_TIMES)
				THEN(*//偏移量为最大的值时,排抓取为最后一排*)
				m_iStep:=5;(*//装盘完成*)
				ELSE
				m_iStep:=2;(*//请求下一次装盘*)			
				IF (m_iCoordinateX-1)/GET_QUANTITY+1=ROW_TIMES THEN
 m_iCoordinateX:=1;                                              (*//开始执行下一列*)
 m_iCoordinateY:=m_iCoordinateY+1;
 ELSE
 m_iCoordinateX:=((m_iCoordinateX-1)/GET_QUANTITY+1)*GET_QUANTITY+1;(*//这一列继续往后排*)
				END_IF;
			END_IF;
		END_IF;
	END_IF;
	5: (*//完成*)
	PackCommunicationIO.o_iSinglePackDonePLCPC:=2;
	IF PackCommunicationIO.i_iSinglePackDoneAknPCPLC =2 THEN
		PackCommunicationIO.o_iSinglePackDonePLCPC:=1;
		m_iCoordinateX:=1;
		m_iCoordinateY:=1;
		FanucRobotIO.io_xMutexLock:=0;
	END_IF;
	IF ConveyorIO.xEmpty AND PackCommunicationIO.o_iSinglePackDonePLCPC=1 THEN
		m_iStep:=1;
	END_IF;
END_CASE;
END_FUNCTION_BLOCK

PROGRAM START
IF g_xReset THEN
	SM50:=1;
	ELSE
	SM50:=0;
END_IF;
CASE g_iState OF
	0: (*手动*)
	g_xManual:=1;
	g_xAuto:=0;	
	g_xStackLampAmber:=1;
	g_xStackLampGreen:=0;
	g_xRemoteAuto:=0;
	g_xAutoLamp:=0;
	1:(*自动*)
	g_xManual:=0;
	g_xAuto:=1;
	g_xStackLampGreen:=1;
	g_xStackLampAmber:=0;
	g_xRemoteAuto:=0;
	g_xAutoLamp:=1;
	2:	(*远程自动*)
	g_xRemoteAuto:=1;
	g_xStackLampGreen:=1;
	g_xStackLampAmber:=0;
	g_xAuto:=0;
	g_xManual:=0;
	g_xAutoLamp:=0;
	3:(*自动未启动*)
	g_xRemoteAuto:=1;
	g_xStackLampGreen:=SM412;
	g_xStackLampAmber:=0;
	g_xAuto:=0;
	g_xManual:=0;	
	g_xAutoLamp:=0;
END_CASE;

IF g_xAutoSwitch AND g_xAutoStart  THEN  
	g_iState:=1;
END_IF;

IF g_xAutoSwitch AND (g_iState<>1 OR NOT g_xStop)  THEN  
	g_iState:=3;
END_IF;

g_xStackLampRed:=g_xAlarm AND SM412;
g_xBuzzer:=g_xAlarm AND SM412 AND NOT g_xMute;

IF LDF(TRUE,g_xAlarm) THEN
	g_xMute:=0;
END_IF;

IF NOT g_xAutoSwitch  OR g_xEStop=0 THEN 
	g_iState:=0;
END_IF;
IF g_xRemoteAutoStart THEN
	g_iState:=2;
END_IF;
IF g_xPause AND SM412 THEN
	g_xStackLampGreen:=0;
	g_xStackLampAmber:=0;
END_IF;
END_PROGRAM

PROGRAM ServoScan
VAR
  istep : INT;  (* 扫码步骤 *)
END_VAR
VAR CONSTANT
  ROW : INT := 8;  (* Y轴每个值对应的电池数量 *)
END_VAR
VAR
  ii : INT;
  jj : INT;
  m_xclean : BOOL;  (* 清零 *)
  kk : INT;  (* 错误位 *)
  m_iLampTwinkle : INT;  (* 灯光闪烁次数 *)
  m_tonScanOvertime : TON;  (* 扫码超时 *)
  m_tScanOvertime : TIME;  (* 扫码超时 *)
  m_xScanOvertime : BOOL;  (* 扫码超时 *)
  m_tonScanDelay : TON;  (* 扫码延时 *)
  m_tScanDelay : TIME;
  m_xScanDelay : BOOL;
END_VAR
Y280:=1;
(*当前位置读取*)
DMOVP(SM412,g_diQD75CurrentPos1,g_diQD75LastPos1);(*记录1S前的位置，和现在的位置比较，判断是否需要重新启动*)
DMOVP(SM412,g_diQD75CurrentPos2,g_diQD75LastPos2);(*记录1S前的位置，和现在的位置比较，判断是否需要重新启动*)
DMOVP(SM412,U28\G800,g_diQD75CurrentPos1);(*双字不能:=，只能dmov了*)
DMOVP(SM412,U28\G900,g_diQD75CurrentPos2);(*双字不能:=，只能dmov了*)
(*如果Y有输出，但是电机没走，那可能是定位过程中发了新的指令，就用这个来断一下Y就能恢复动作了*)
IF (g_yQD75LocateStart1 AND g_diQD75CurrentPos1=g_diQD75LastPos1 )
	 OR (g_yQD75LocateStart2 AND g_diQD75CurrentPos2=g_diQD75LastPos2 ) THEN
				g_xResetServo:=1;
ELSE
				g_xResetServo:=0;
END_IF;		
(*目标地址读取*)
g_iQD75LastNumber1:=U28\G837;(*上一次目标号*)
g_iQD75DestiNumber1:=U28\G835;(*目标号*)
DMOV(TRUE,U28\G818,g_diQD75DestinationPos1);(*目标地址*)
g_iQD75LastNumber2:=U28\G937;(*上一次目标号*)
g_iQD75DestiNumber2:=U28\G935;(*目标号*)
DMOV(TRUE,U28\G918,g_diQD75DestinationPos2);(*目标地址*)
(*报警信息读取*)
g_iQD75ErrorNumber1:=U28\G806;
g_iQD75ErrorNumber2:=U28\G906;
(*报警复位*)
IF LDP(TRUE,g_xResetServo) THEN
	U28\G1502:=1;(*X轴复位*)(*这俩信号都能自动复位*)
	U28\G1602:=1;(*Y轴复位*)
	U28\G1503:=1;(*X轴重起*)
	U28\G1603:=1;(*Y轴重起*)
	(*YBE:= X78 OR  X79;*)(*X78,X79为两个驱动器的报警，这个驱动器只能断电复位，所以YAE控制断电*)
(*ELSE
	YBE:=0*);
	
END_IF;	







(*下面是正式流程*)
(*除了正常运过去那种，有时手动放上去的也要能启动扫码流程，要加个按钮*)
SET( g_xPutInto, g_xServoStart );
 CASE istep OF 
 0:(*初始化，等待启动信号*)
 				U28\G1500:=9001;(*9001表示会回原点*)
 				U28\G1600:=9001;
 				g_yQD75LocateStart1:= NOT g_xResetServo AND NOT g_xQD75LocateDone1
 																AND U28\G800<>0;
 				g_yQD75LocateStart2:= NOT g_xResetServo AND NOT g_xQD75LocateDone2
 																AND U28\G900<>0;		
 				MOV( g_xServoStart AND U28\G800=0 AND U28\G900=0, 10, istep );(*800是当前位置值*)
 	(*10是在0之后，1之前的一个步骤，扫框码，等待扫码完成。懒得改，就插在这里了*)
 10:(*扫框码，扫码完成再去扫电池码*)
 				(*夹紧气缸夹住*)
 				g_yQD75LocateStart1:=0;
 				g_yQD75LocateStart2:=0;
 				g_xCatchCylinder:=1;
 	 			g_xServoStart:=0;
 				g_xScan:=0; 	
 				D3000:=2;(**扫框码请求**)
 				IF D2000=2 THEN(*扫码成功*)
 							g_iXaxisNumber:=1;
 							g_iYaxisNumber:=1;
 							istep:=1;
 				END_IF;	
 1:(*伺服行走*)
 				(*X轴行走*)	
 				IF NOT g_xQD75LocateDone1 AND g_iXaxisNumber<>0 THEN(*起始地址设定是100，那么g_xQD75LocateDone1就是1轴定位完成信号*)
 							U28\G1500:=g_iXaxisNumber;(*起始地址设定是100，这里就要写U28，起始地址去掉个0。G1500是X轴定位启动的编号*)
 							g_yQD75LocateStart1:=NOT g_xQD75Error1;(*起始地址设定是100，那么g_yQD75LocateStart1就是1轴定位启动信号*)
 				ELSE
 							U28\G1500:=0;
 							g_yQD75LocateStart1:=0;
 				END_IF;		
 				(*Y轴行走*)	
 				IF NOT g_xQD75LocateDone2 AND g_iYaxisNumber<>0 THEN
 							U28\G1600:=g_iYaxisNumber;
 							g_yQD75LocateStart2:=NOT g_xQD75Error2;
 				ELSE
 							U28\G1600:=0;
 							g_yQD75LocateStart2:=0;
 				END_IF;	
 				SET( g_xQD75LocateDone1 AND g_xQD75LocateDone2 , g_xScan);
 				MOV( g_xQD75LocateDone1 AND g_xQD75LocateDone2 , 2, istep );
 2:(*进行扫码*)
 				g_yQD75LocateStart1:=0;
 				g_yQD75LocateStart2:=0;
 				(*扫码结果为8，表示扫码错误，调回step1，重新扫一次*)
 				IF g_iBatteryInformation[0]=8 AND TS63 THEN
 							g_iBatteryInformation[0]:=0;
 							g_xScan:=0;(*_
 							IF  g_iXaxisNumber<20 THEN_*)(*表示第一次扫码尝试失败*)(*_
 										g_iXaxisNumber:=g_iXaxisNumber+20;
 										g_iYaxisNumber:=g_iYaxisNumber+20;
 										istep:=1;
 							ELSIF g_iXaxisNumber>20 THEN_*)(*表示第二次扫码失败，两次都扫失败就跳过了*)
 										FOR ii:=0 TO 10 DO
 													IF g_iScanError[ii]=0 THEN(*把错误字都存起来，完成任务清零*)
 															g_iScanError[ii]:=g_iBatteryPosition;
 															g_iErrorSUM:=ii+1;
 															EXIT;
 													END_IF;
 										END_FOR;	
 											
 										IF g_iBatteryPosition>0 AND g_iBatteryPosition<128 AND TS63 THEN
 										(*数据复位*)
 													FOR jj:=0 TO 16 DO
 															g_iBatteryInformation[jj]:=0;
 													END_FOR;
 										(*这里的框是特殊形状的，有16列，每列对应8排，但是基数列和偶数列又是错开的，所以单独写的位置计算*)
 				 									g_iBatteryPosition:=g_iBatteryPosition+1;
 													g_iXaxisNumber:=(g_iBatteryPosition-1)/ROW+1;
 													g_iYaxisNumber:=2*((g_iBatteryPosition-1)MOD ROW)+1+((g_iXaxisNumber-1) MOD 2);(*后面这个是判断奇偶的，奇数列不加，偶数列加1*)
 													istep:=1;
 										ELSIF g_iBatteryPosition=128 AND TS63 THEN
 													FOR jj:=0 TO 16 DO
 																g_iBatteryInformation[jj]:=0;
 													END_FOR;
 													istep:=3;	
 										END_IF;			
 							(*_END_IF;	_*)
 				END_IF;	
 				Z0:=(g_iBatteryPosition-1)*15;(*正常情况，每个电池占用15个字,-1是因为位置参数是从1开始，不是0开始*)
 				IF g_xScan AND g_iBatteryInformation[0]=24 THEN(*扫码成功会有24个字，不成功会有8个字，还可能读错，就会超过24个字，都属于不正常*)
 							D3006Z0:=g_iBatteryInformation[1];
 							D3007Z0:=g_iBatteryInformation[2];(*1-14都是电池码*)
 							D3008Z0:=g_iBatteryInformation[3];
 							D3009Z0:=g_iBatteryInformation[4];
 							D3010Z0:=g_iBatteryInformation[5];
 							D3011Z0:=g_iBatteryInformation[6];
 							D3012Z0:=g_iBatteryInformation[7];
 							D3013Z0:=g_iBatteryInformation[8];
 							D3014Z0:=g_iBatteryInformation[9];
 							D3015Z0:=g_iBatteryInformation[10];
 							D3016Z0:=g_iBatteryInformation[11];
 							D3017Z0:=g_iBatteryInformation[12];
 							D3018Z0:=g_iBatteryInformation[13];
 							D3019Z0:=g_iBatteryInformation[14];
 							D3020Z0:=g_iBatteryInformation[15];
 							IF g_iBatteryPosition>0 AND g_iBatteryPosition<128 AND TS63 THEN
 										g_xScan:=0;
 										(*数据复位*)
 										FOR jj:=0 TO 16 DO
 													g_iBatteryInformation[jj]:=0;
 										END_FOR;
 										(*这里的框是特殊形状的，有16列，每列对应8排，但是基数列和偶数列又是错开的，所以单独写的位置计算*)
 				 						g_iBatteryPosition:=g_iBatteryPosition+1;
 										g_iXaxisNumber:=(g_iBatteryPosition-1)/ROW+1;
 										g_iYaxisNumber:=2*((g_iBatteryPosition-1)MOD ROW)+1+((g_iXaxisNumber-1) MOD 2);(*后面这个是判断奇偶的，奇数列不加，偶数列加1*)
 										istep:=1;
 						ELSIF g_iBatteryPosition=128 AND TS63 THEN
 										FOR jj:=0 TO 16 DO
 													g_iBatteryInformation[jj]:=0;
 										END_FOR;
 										g_xScan:=0;
 										istep:=3;	
 						END_IF;(*位置在1-128之间那个if*)
 				END_IF;(*扫码成功那个if*)		
 3:(*数据上传*)
   				IF g_iScanError[6]=0 THEN
 							D3001:=2;(*装载完成，数据上传*)
 				END_IF;
 				IF D2001=2 THEN(*表示数据收到，可以放行*)
 							istep:=4;
 				END_IF;
 4:(*数据复位，下料，回0步*)
 				D3001:=1;
 				g_xCatchCylinder:=0;
 				g_xScanDone:=1;
 				IF X280 THEN
 							U28\G1500:=1;
 							U28\G1600:=1;
 							g_yQD75LocateStart1:=NOT g_xQD75LocateDone1 AND NOT g_xQD75Error1;
 							g_yQD75LocateStart2:=NOT g_xQD75LocateDone2 AND NOT g_xQD75Error2;
 				END_IF;
 20:(*这里加一个专门去不良位的，调试用*)
 				 D2009:=g_iScanError[0]+g_iScanError[1](*这个没有意义，只是为了方便我看没扫上的那些位置*)
 								+g_iScanError[2]+g_iScanError[3]+g_iScanError[ 4]
								+g_iScanError[5] +g_iScanError[6] +g_iScanError[7]
  								+g_iScanError[8]+g_iScanError[9];
 				g_iXaxisNumber:=(kk-1)/ROW+1;
 				g_iYaxisNumber:=2*((kk-1)MOD ROW)+1+((g_iXaxisNumber-1) MOD 2);
 				U28\G1500:=g_iXaxisNumber;
 				U28\G1600:=g_iYaxisNumber; 
 				DMOV(TRUE,10000,U28\G1518);
 				DMOV(TRUE,10000,U28\G1618);
 				g_yQD75LocateStart1:=NOT g_xQD75LocateDone1 AND NOT g_yQD75JogCW1 AND NOT g_yQD75JogCCW1 AND NOT g_xQD75Error1;
 				g_yQD75LocateStart2:=NOT g_xQD75LocateDone2 AND NOT g_yQD75JogCW2 AND NOT g_yQD75JogCCW2 AND NOT g_xQD75Error1;
 				g_yQD75JogCW1:=NOT g_yQD75JogCCW1 AND g_xJogXCW;(*1轴JOG正转*)
 				g_yQD75JogCCW1:=NOT g_yQD75JogCW1 AND g_xJogXCCW;(*1轴JOG反转*)
 				g_yQD75JogCW2:=NOT g_yQD75JogCCW2 AND g_xJogYCW;(*2轴JOG正转*)
 				g_yQD75JogCCW2:=NOT g_yQD75JogCW2 AND g_xJogYCCW;(*2轴JOG反转*)
 				
 END_CASE;
(*这个写在case外边，方便复位*) 
IF TS60 AND NOT g_xQD75Busy1 AND NOT g_xQD75Busy2 THEN
	(*T190是下料时，离开开关延时，离开开关这么久就认为物料已远走，可以开始运下一个了*)
 			FOR Z1:=0 TO 1920 DO(*物料送走，数据复位*)
 						D3006Z1:=0;
 		 	END_FOR;
 		  	D3000:=1;(*扫框码请求复位*)
 		  	g_xServoStart:=0;
 			g_xScanDone:=0;
 			g_iBatteryPosition:=1;
 			istep:=0;
END_IF;
 m_tonScanDelay(IN:=g_iBatteryInformation[0]<>0 AND istep=2,PT:=t#100ms,Q:= m_xScanDelay ,ET:= m_tScanDelay);;(*扫码成功到接收数据完毕需要时间，所以做个延时*)
 OUT_T( g_iBatteryInformation[0]<>0 AND istep=2 , TC63 ,k3 );
 m_tonScanOvertime(IN:=g_iBatteryInformation[0]=0 AND istep=2 AND NOT g_xScanOvertime  ,PT:=t#1S ,Q:= g_xScanOvertime ,ET:= m_tScanOvertime );(*有时候扫码请求发出去数据没接收到，需要重新启动扫码，等10S*)
 IF TS60 OR m_xclean THEN
 	FOR jj:=0 TO 9 DO
 		g_iScanError[jj]:=0;
 	END_FOR;
 	g_iErrorSUM:=0;
 END_IF;		
 YBA:=g_iScanError[5]<>0;(*超过6个就报警,而且放行*)
 (*IF ldp(TRUE,g_iScanError[5]<>0 )THEN
 		g_xScanDone:=1;
 END_IF;	*)
END_PROGRAM
